TYPE UDT_MAN_CMD_WR :   // Manual commands from HMI
STRUCT
   CONV_Manual_ALL : BOOL;
   CONV_Man_ALL_FWD : BOOL;
   CONV_Man_ALL_REV : BOOL;
   M302M1_Manual : BOOL;
   M302M1_ManFWD : BOOL;
   M302M1_ManREV : BOOL;
   M302M1_ManSpeed : DINT;
   M302M2_Manual : BOOL;
   M302M2_ManFWD : BOOL;
   M302M2_ManREV : BOOL;
   M302M2_ManSpeed : DINT;
   M302M3_Manual : BOOL;
   M302M3_ManFWD : BOOL;
   M302M3_ManREV : BOOL;
   M302M3_ManSpeed : DINT;
   M302M4_Manual : BOOL;
   M302M4_ManFWD : BOOL;
   M302M4_ManREV : BOOL;
   M302M4_ManSpeed : DINT;
   M302M5_Manual : BOOL;
   M302M5_ManFWD : BOOL;
   M302M5_ManREV : BOOL;
   M302M5_ManSpeed : DINT;
   M302M6_Manual : BOOL;
   M302M6_ManFWD : BOOL;
   M302M6_ManREV : BOOL;
   M302M6_ManSpeed : DINT;
   M302M7_Manual : BOOL;
   M302M7_ManFWD : BOOL;
   M302M7_ManREV : BOOL;
   M302M7_ManSpeed : DINT;
   M303M1_Manual : BOOL;
   M303M1_ManFWD : BOOL;
   M303M1_ManREV : BOOL;
   M303M1_ManSpeed : DINT;
   M303M2_Manual : BOOL;
   M303M2_ManFWD : BOOL;
   M303M2_ManREV : BOOL;
   M303M2_ManSpeed : DINT;
   M304M1_Manual : BOOL;
   M304M1_ManFWD : BOOL;
   M304M1_ManREV : BOOL;
   M304M1_ManSpeed : DINT;
   M305M1_Manual : BOOL;
   M305M1_ManFWD : BOOL;
   M305M1_ManREV : BOOL;
   M305M1_ManSpeed : DINT;
   M306M1_Manual : BOOL;
   M306M1_ManFWD : BOOL;
   M306M1_ManREV : BOOL;
   M306M1_ManSpeed : DINT;
   M307AM1_Manual : BOOL;
   M307AM1_ManFWD : BOOL;
   M307AM1_ManREV : BOOL;
   M307AM1_ManSpeed : DINT;
   M307AM2_Manual : BOOL;
   M307AM2_ManFWD : BOOL;
   M307AM2_ManREV : BOOL;
   M307AM2_ManSpeed : DINT;
   M307AM3_Manual : BOOL;
   M307AM3_ManFWD : BOOL;
   M307AM3_ManREV : BOOL;
   M307AM3_ManSpeed : DINT;
   M307AM4_Manual : BOOL;
   M307AM4_ManFWD : BOOL;
   M307AM4_ManREV : BOOL;
   M307AM4_ManSpeed : DINT;
   M307BM1_Manual : BOOL;
   M307BM1_ManFWD : BOOL;
   M307BM1_ManREV : BOOL;
   M307BM1_ManSpeed : DINT;
   M307CM1_Manual : BOOL;
   M307CM1_ManFWD : BOOL;
   M307CM1_ManREV : BOOL;
   M307CM1_ManSpeed : DINT;
   M307DM1_Manual : BOOL;
   M307DM1_ManFWD : BOOL;
   M307DM1_ManREV : BOOL;
   M307DM1_ManSpeed : DINT;
   M307EM1_Manual : BOOL;
   M307EM1_ManFWD : BOOL;
   M307EM1_ManREV : BOOL;
   M307EM1_ManSpeed : DINT;
   M307FM1_Manual : BOOL;
   M307FM1_ManFWD : BOOL;
   M307FM1_ManREV : BOOL;
   M307FM1_ManSpeed : DINT;
   M310M1_Manual : BOOL;
   M310M1_ManFWD : BOOL;
   M310M1_ManREV : BOOL;
   M310M1_ManSpeed : DINT;
   M310M2_Manual : BOOL;
   M310M2_ManFWD : BOOL;
   M310M2_ManREV : BOOL;
   M310M2_ManSpeed : DINT;
   M310M3_Manual : BOOL;
   M310M3_ManFWD : BOOL;
   M310M3_ManREV : BOOL;
   M310M3_ManSpeed : DINT;
   M310M4_Manual : BOOL;
   M310M4_ManFWD : BOOL;
   M310M4_ManREV : BOOL;
   M310M4_ManSpeed : DINT;
   M310M5_Manual : BOOL;
   M310M5_ManFWD : BOOL;
   M310M5_ManREV : BOOL;
   M310M5_ManSpeed : DINT;
   M310M6_Manual : BOOL;
   M310M6_ManFWD : BOOL;
   M310M6_ManREV : BOOL;
   M310M6_ManSpeed : DINT;
   M310M7_Manual : BOOL;
   M310M7_ManFWD : BOOL;
   M310M7_ManREV : BOOL;
   M310M7_ManSpeed : DINT;
   M311M1_Manual : BOOL;
   M311M1_ManFWD : BOOL;
   M311M1_ManREV : BOOL;
   M311M1_ManSpeed : DINT;
   M311AM1_Manual : BOOL;
   M311AM1_ManFWD : BOOL;
   M311AM1_ManREV : BOOL;
   M311AM1_ManSpeed : DINT;
   M312M1_Manual : BOOL;
   M312M1_ManFWD : BOOL;
   M312M1_ManREV : BOOL;
   M312M1_ManSpeed : DINT;
   M312M2_Manual : BOOL;
   M312M2_ManFWD : BOOL;
   M312M2_ManREV : BOOL;
   M312M2_ManSpeed : DINT;
   M312M3_Manual : BOOL;
   M312M3_ManFWD : BOOL;
   M312M3_ManREV : BOOL;
   M312M3_ManSpeed : DINT;
   M315M1_Manual : BOOL;
   M315M1_ManFWD : BOOL;
   M315M1_ManREV : BOOL;
   M315M1_ManSpeed : DINT;
   M315M2_Manual : BOOL;
   M315M2_ManFWD : BOOL;
   M315M2_ManREV : BOOL;
   M315M2_ManSpeed : DINT;
   M315M3_Manual : BOOL;
   M315M3_ManFWD : BOOL;
   M315M3_ManREV : BOOL;
   M315M3_ManSpeed : DINT;
   M315M4_Manual : BOOL;
   M315M4_ManFWD : BOOL;
   M315M4_ManREV : BOOL;
   M315M4_ManSpeed : DINT;
   M315M5_Manual : BOOL;
   M315M5_ManFWD : BOOL;
   M315M5_ManREV : BOOL;
   M315M5_ManSpeed : DINT;
   M315M6_Manual : BOOL;
   M315M6_ManFWD : BOOL;
   M315M6_ManREV : BOOL;
   M315M6_ManSpeed : DINT;
   M315M7_Manual : BOOL;
   M315M7_ManFWD : BOOL;
   M315M7_ManREV : BOOL;
   M315M7_ManSpeed : DINT;
   M315AM1_Manual : BOOL;
   M315AM1_ManFWD : BOOL;
   M315AM1_ManREV : BOOL;
   M315AM1_ManSpeed : DINT;
   M316M1_Manual : BOOL;
   M316M1_ManFWD : BOOL;
   M316M1_ManREV : BOOL;
   M316M1_ManSpeed : DINT;
   M316AM1_Manual : BOOL;
   M316AM1_ManFWD : BOOL;
   M316AM1_ManREV : BOOL;
   M316AM1_ManSpeed : DINT;
   M317M1_Manual : BOOL;
   M317M1_ManFWD : BOOL;
   M317M1_ManREV : BOOL;
   M317M1_ManSpeed : DINT;
   M317M2_Manual : BOOL;
   M317M2_ManFWD : BOOL;
   M317M2_ManREV : BOOL;
   M317M2_ManSpeed : DINT;
   M317M3_Manual : BOOL;
   M317M3_ManFWD : BOOL;
   M317M3_ManREV : BOOL;
   M317M3_ManSpeed : DINT;
   M350M1_Manual : BOOL;
   M350M1_ManFWD : BOOL;
   M350M1_ManREV : BOOL;
   M350M1_ManSpeed : DINT;
   M351M1_Manual : BOOL;
   M351M1_ManFWD : BOOL;
   M351M1_ManREV : BOOL;
   M351M1_ManSpeed : DINT;
   M360M1_Manual : BOOL;
   M360M1_ManFWD : BOOL;
   M360M1_ManREV : BOOL;
   M360M1_ManSpeed : DINT;
END_STRUCT
END_TYPE

TYPE UDT_MOTOR_HMR :
STRUCT
   M302M1_Feedback : BOOL;
   M302M1_Faulted : BOOL;
   M302M1_FaultCode : DINT;
   M302M1_OutSpeed : DINT;
   M302M1_OutCurrent : DINT;
   M302M2_Feedback : BOOL;
   M302M2_Faulted : BOOL;
   M302M2_FaultCode : DINT;
   M302M2_OutSpeed : DINT;
   M302M2_OutCurrent : DINT;
   M302M3_Feedback : BOOL;
   M302M3_Faulted : BOOL;
   M302M3_FaultCode : DINT;
   M302M3_OutSpeed : DINT;
   M302M3_OutCurrent : DINT;
   M302M4_Feedback : BOOL;
   M302M4_Faulted : BOOL;
   M302M4_FaultCode : DINT;
   M302M4_OutSpeed : DINT;
   M302M4_OutCurrent : DINT;
   M302M5_Feedback : BOOL;
   M302M5_Faulted : BOOL;
   M302M5_FaultCode : DINT;
   M302M5_OutSpeed : DINT;
   M302M5_OutCurrent : DINT;
   M302M6_Feedback : BOOL;
   M302M6_Faulted : BOOL;
   M302M6_FaultCode : DINT;
   M302M6_OutSpeed : DINT;
   M302M6_OutCurrent : DINT;
   M302M7_Feedback : BOOL;
   M302M7_Faulted : BOOL;
   M302M7_FaultCode : DINT;
   M302M7_OutSpeed : DINT;
   M302M7_OutCurrent : DINT;
   M303M1_Feedback : BOOL;
   M303M1_Faulted : BOOL;
   M303M1_FaultCode : DINT;
   M303M1_OutSpeed : DINT;
   M303M1_OutCurrent : DINT;
   M303M2_Feedback : BOOL;
   M303M2_Faulted : BOOL;
   M303M2_FaultCode : DINT;
   M303M2_OutSpeed : DINT;
   M303M2_OutCurrent : DINT;
   M304M1_Feedback : BOOL;
   M304M1_Faulted : BOOL;
   M304M1_FaultCode : DINT;
   M304M1_OutSpeed : DINT;
   M304M1_OutCurrent : DINT;
   M305M1_Feedback : BOOL;
   M305M1_Faulted : BOOL;
   M305M1_FaultCode : DINT;
   M305M1_OutSpeed : DINT;
   M305M1_OutCurrent : DINT;
   M306M1_Feedback : BOOL;
   M306M1_Faulted : BOOL;
   M306M1_FaultCode : DINT;
   M306M1_OutSpeed : DINT;
   M306M1_OutCurrent : DINT;
   M307AM1_Feedback : BOOL;
   M307AM1_Faulted : BOOL;
   M307AM1_FaultCode : DINT;
   M307AM1_OutSpeed : DINT;
   M307AM1_OutCurrent : DINT;
   M307AM2_Feedback : BOOL;
   M307AM2_Faulted : BOOL;
   M307AM2_FaultCode : DINT;
   M307AM2_OutSpeed : DINT;
   M307AM2_OutCurrent : DINT;
   M307AM3_Feedback : BOOL;
   M307AM3_Faulted : BOOL;
   M307AM3_FaultCode : DINT;
   M307AM3_OutSpeed : DINT;
   M307AM3_OutCurrent : DINT;
   M307AM4_Feedback : BOOL;
   M307AM4_Faulted : BOOL;
   M307AM4_FaultCode : DINT;
   M307AM4_OutSpeed : DINT;
   M307AM4_OutCurrent : DINT;
   M307BM1_Feedback : BOOL;
   M307BM1_Faulted : BOOL;
   M307BM1_FaultCode : DINT;
   M307BM1_OutSpeed : DINT;
   M307BM1_OutCurrent : DINT;
   M307CM1_Feedback : BOOL;
   M307CM1_Faulted : BOOL;
   M307CM1_FaultCode : DINT;
   M307CM1_OutSpeed : DINT;
   M307CM1_OutCurrent : DINT;
   M307DM1_Feedback : BOOL;
   M307DM1_Faulted : BOOL;
   M307DM1_FaultCode : DINT;
   M307DM1_OutSpeed : DINT;
   M307DM1_OutCurrent : DINT;
   M307EM1_Feedback : BOOL;
   M307EM1_Faulted : BOOL;
   M307EM1_FaultCode : DINT;
   M307EM1_OutSpeed : DINT;
   M307EM1_OutCurrent : DINT;
   M307FM1_Feedback : BOOL;
   M307FM1_Faulted : BOOL;
   M307FM1_FaultCode : DINT;
   M307FM1_OutSpeed : DINT;
   M307FM1_OutCurrent : DINT;
   M310M1_Feedback : BOOL;
   M310M1_Faulted : BOOL;
   M310M1_FaultCode : DINT;
   M310M1_OutSpeed : DINT;
   M310M1_OutCurrent : DINT;
   M310M2_Feedback : BOOL;
   M310M2_Faulted : BOOL;
   M310M2_FaultCode : DINT;
   M310M2_OutSpeed : DINT;
   M310M2_OutCurrent : DINT;
   M310M3_Feedback : BOOL;
   M310M3_Faulted : BOOL;
   M310M3_FaultCode : DINT;
   M310M3_OutSpeed : DINT;
   M310M3_OutCurrent : DINT;
   M310M4_Feedback : BOOL;
   M310M4_Faulted : BOOL;
   M310M4_FaultCode : DINT;
   M310M4_OutSpeed : DINT;
   M310M4_OutCurrent : DINT;
   M310M5_Feedback : BOOL;
   M310M5_Faulted : BOOL;
   M310M5_FaultCode : DINT;
   M310M5_OutSpeed : DINT;
   M310M5_OutCurrent : DINT;
   M310M6_Feedback : BOOL;
   M310M6_Faulted : BOOL;
   M310M6_FaultCode : DINT;
   M310M6_OutSpeed : DINT;
   M310M6_OutCurrent : DINT;
   M310M7_Feedback : BOOL;
   M310M7_Faulted : BOOL;
   M310M7_FaultCode : DINT;
   M310M7_OutSpeed : DINT;
   M310M7_OutCurrent : DINT;
   M311M1_Feedback : BOOL;
   M311M1_Faulted : BOOL;
   M311M1_FaultCode : DINT;
   M311M1_OutSpeed : DINT;
   M311M1_OutCurrent : DINT;
   M311AM1_Feedback : BOOL;
   M311AM1_Faulted : BOOL;
   M311AM1_FaultCode : DINT;
   M311AM1_OutSpeed : DINT;
   M311AM1_OutCurrent : DINT;
   M312M1_Feedback : BOOL;
   M312M1_Faulted : BOOL;
   M312M1_FaultCode : DINT;
   M312M1_OutSpeed : DINT;
   M312M1_OutCurrent : DINT;
   M312M2_Feedback : BOOL;
   M312M2_Faulted : BOOL;
   M312M2_FaultCode : DINT;
   M312M2_OutSpeed : DINT;
   M312M2_OutCurrent : DINT;
   M312M3_Feedback : BOOL;
   M312M3_Faulted : BOOL;
   M312M3_FaultCode : DINT;
   M312M3_OutSpeed : DINT;
   M312M3_OutCurrent : DINT;
   M315M1_Feedback : BOOL;
   M315M1_Faulted : BOOL;
   M315M1_FaultCode : DINT;
   M315M1_OutSpeed : DINT;
   M315M1_OutCurrent : DINT;
   M315M2_Feedback : BOOL;
   M315M2_Faulted : BOOL;
   M315M2_FaultCode : DINT;
   M315M2_OutSpeed : DINT;
   M315M2_OutCurrent : DINT;
   M315M3_Feedback : BOOL;
   M315M3_Faulted : BOOL;
   M315M3_FaultCode : DINT;
   M315M3_OutSpeed : DINT;
   M315M3_OutCurrent : DINT;
   M315M4_Feedback : BOOL;
   M315M4_Faulted : BOOL;
   M315M4_FaultCode : DINT;
   M315M4_OutSpeed : DINT;
   M315M4_OutCurrent : DINT;
   M315M5_Feedback : BOOL;
   M315M5_Faulted : BOOL;
   M315M5_FaultCode : DINT;
   M315M5_OutSpeed : DINT;
   M315M5_OutCurrent : DINT;
   M315M6_Feedback : BOOL;
   M315M6_Faulted : BOOL;
   M315M6_FaultCode : DINT;
   M315M6_OutSpeed : DINT;
   M315M6_OutCurrent : DINT;
   M315M7_Feedback : BOOL;
   M315M7_Faulted : BOOL;
   M315M7_FaultCode : DINT;
   M315M7_OutSpeed : DINT;
   M315M7_OutCurrent : DINT;
   M315AM1_Feedback : BOOL;
   M315AM1_Faulted : BOOL;
   M315AM1_FaultCode : DINT;
   M315AM1_OutSpeed : DINT;
   M315AM1_OutCurrent : DINT;
   M316M1_Feedback : BOOL;
   M316M1_Faulted : BOOL;
   M316M1_FaultCode : DINT;
   M316M1_OutSpeed : DINT;
   M316M1_OutCurrent : DINT;
   M316AM1_Feedback : BOOL;
   M316AM1_Faulted : BOOL;
   M316AM1_FaultCode : DINT;
   M316AM1_OutSpeed : DINT;
   M316AM1_OutCurrent : DINT;
   M317M1_Feedback : BOOL;
   M317M1_Faulted : BOOL;
   M317M1_FaultCode : DINT;
   M317M1_OutSpeed : DINT;
   M317M1_OutCurrent : DINT;
   M317M2_Feedback : BOOL;
   M317M2_Faulted : BOOL;
   M317M2_FaultCode : DINT;
   M317M2_OutSpeed : DINT;
   M317M2_OutCurrent : DINT;
   M317M3_Feedback : BOOL;
   M317M3_Faulted : BOOL;
   M317M3_FaultCode : DINT;
   M317M3_OutSpeed : DINT;
   M317M3_OutCurrent : DINT;
   M350M1_Feedback : BOOL;
   M350M1_Faulted : BOOL;
   M350M1_FaultCode : DINT;
   M350M1_OutSpeed : DINT;
   M350M1_OutCurrent : DINT;
   M351M1_Feedback : BOOL;
   M351M1_Faulted : BOOL;
   M351M1_FaultCode : DINT;
   M351M1_OutSpeed : DINT;
   M351M1_OutCurrent : DINT;
   M360M1_Feedback : BOOL;
   M360M1_Faulted : BOOL;
   M360M1_FaultCode : DINT;
   M360M1_OutSpeed : DINT;
   M360M1_OutCurrent : DINT;
END_STRUCT
END_TYPE

TYPE UDT_PLANT_CONSTANTS :
STRUCT
   dPLC_ID : DINT;   // 1= PLC#1 2= PLC#2
   dOP_Side : DINT;   // 0=Operator side right; 1=Operator side left
   dZ1ConveyorNumber : DINT;   // Conveyor number in Z301
   dZ1TotalLength_cmm : DINT;   // Z301 total length of tracking [mm/100]
   dZ2ConveyorNumber : DINT;   // Conveyor number in Z302
   dZ2TotalLength_cmm : DINT;   // Z302 total length of tracking [mm/100]
   dZ3ConveyorNumber : DINT;   // Conveyor number in Z303
   dZ3TotalLength_cmm : DINT;   // Z303 total length of tracking [mm/100]
   dTrimDeckNumber : DINT;   // Trimming deck number
   dTrimWheelsNumber : DINT;   // Trimming wheels number
   dSplitBarNumber : DINT;   // Split bar number
   dSepRollNumber : DINT;   // Separator roll number
   dTrackWindows_cmm : DINT;   // Tracking windows step [mm/100]
   dMaxScanSpace_cmm : DINT;   // Max space calculated on each scan at maximum line speed [mm/100]
   rgdAccDecRamps : REAL[4];   // Acceleration / Deceleration ramps used in main line [m/s2]
   dMaxLineSpeed_mm_min : DINT;   // Max line speed [mm/min]
   dMinLineSpeed_mm_min : DINT;   // Min line speed [mm/min]
   dMaxLineSnapSpeed_mm_min : DINT;   // Max line speed for snapping area [mm/min]
   dMinLineSnapSpeed_mm_min : DINT;   // Min line speed for snapping area [mm/min]
   dMaxLehrSpeed_mm_min : DINT;   // Max lehr speed [mm/min]
   dMinLehrSpeed_mm_min : DINT;   // Min lehr speed [mm/min]
   rMaxSpeedRatio : REAL;   // Max speed ratio [Num]
   rMinSpeedRatio : REAL;   // Min speed ratio [Num]
   rMaxSpeedSnapRatio : REAL;   // Max speed ratio for snapping area [Num]
   rMinSpeedSnapRatio : REAL;   // Min speed ratio for snapping area [Num]
   dZ1CleaningSpeed_mm_min : DINT;   // Cleaning speed Z301 [mm/min] (Optional if no cooling on motors)
   dMaxNumPlates : DINT;   // Maximum number of plates in tracking (circular buffer positions)
   dMaxNumHeadTail : DINT;   // Maximum number of head tail
   rgdLiteLimits_cmm : DINT[20];   // Lite limits [mm/100] (Length,width...)
   rgdCapLimits_cmm : DINT[5];   // Cap limits [mm/100] (Length,width,max num lites,...)
   rgdConvoyLimits_cmm : DINT[5];   // Convoy limits [mm/100] (Length,width,max num caps,...)
   rgdRibbonLimits_cmm : DINT[5];   // Ribbon limits [mm/100]
   rgdWanderLimits : DINT[2];   // Wander limits [mm/100]
   dNumOfConveyors : DINT;   // Number of conveyors [Num]
   dNumCapsConveyor : DINT;   // Number of caps per conveyor [Num]
   dNumCapsMaxConvoy : DINT;   // Maximum number of caps per convoy [Num]
   dNumLitesMaxCap : DINT;   // Maximum number of lites per cap [Num]
   dNumPlateSearch : DINT;   // Number of plates to search in Search function [Num]
   dNumOfUnloadDestinations : DINT;   // Number of possible destinations for stack [Num]
END_STRUCT
END_TYPE

TYPE UDT_PlateData_Convoy :
STRUCT
   dSyncHead : DINT;   // Synchro Head
   dIDTx : DINT;
   dTotLenght_cmm : DINT;
   dTotWidth_cmm : DINT;
   dFormat : DINT;   // 1=JS 2=LES, 3=SSS
   dNumLites : DINT;   // Num Lite on board
   dPositionLite : DINT;   // 0=Centre Line, 1=Right Side Line. 2 Left Side Line
   tLite : UDT_PlateData_Convoy_Lite[2];
   dSyncTail : DINT;   // Synchro Tail
END_STRUCT
END_TYPE

TYPE UDT_PlateData_Convoy_Lite :
STRUCT
   dID : DINT;   // ID lite
   dProduction_ID : DINT;   // ID Production
   dLenght_cmm : DINT;   // Lenght Lite
   dWidth_cmm : DINT;   // Width Lite
   dThick_cmm : DINT;   // Thickness Lite
   rgxOrigin : DINT;   // Origin plate
   rgxMain : DINT;   // Main destination plate
   rgxAlternative : DINT;   // Alternative destination plate
   xCoated : BOOL;   // Type Coated
   xCoverPlate : BOOL;   // Type Cover
END_STRUCT
END_TYPE

TYPE UDT_SearchPlateAuxData :   // Auxiliary data for searching plate
STRUCT
   dIDMemory : DINT;   // ID Memory
   dReaction_cmm : DINT;   // Reation space [mm/100]
   dPositionDecision_cmm : DINT;   // Decision position [mm/100]
   dPositionStopSearch_cmm : DINT;   // Stop search position [mm/100]
   dPositionStopHooked_cmm : DINT;   // Stop hooked position [mm/100]
   dIndex : DINT;   // Index
   xIndexCons : BOOL;   // Index consistent
   xPlateHooked : BOOL;   // Plate hooked
   OS_xPlateInWindows : BOOL;   // OS Plate in windows
   OF_xPlateInWindows : BOOL;   // OF Plate in windows
   OSR_xPlateInWindows : BOOL;   // OSR Plate in windows
   OSF_xPlateInWindows : BOOL;   // OSF Plate in windows
   OSR_xPlateOutHooked : BOOL;   // OSR Plate hooked
   OS_xPlateOutHooked : BOOL;   // OS Plate hooked
   tResult : GP_TrackingSearchPlate_STC;   // Search plate data result
END_STRUCT
END_TYPE

TYPE UDT_StandConv :
STRUCT
   ST_rgxRampInProgress : DINT;   // Ramp in progress
   ST_rgxDecInProgress : DINT;   // Deceleration in progress
   ST_rgxAccInProgress : DINT;   // Acceleration in progress
   ST_rgxBrakeRelease : DINT;   // Brake release
   ST_rgxBrakeFeedback : DINT;   // Brake feedback
   ST_rgxConveyorOutRunSgm : DINT;   // Single motor conveyor out run
   ST_rgxOutMotorRunSgm : DINT;   // Single motor out run active
   ST_xDriveInDec : BOOL;   // At least one drive in deceleration
   ST_xPositionReached : BOOL;   // Position reached
   ST_xManualCmdEnabled : BOOL;   // Manual command enabled
   ST_xEnableControlError : BOOL;   // Enable control error
   ST_xRotationFeedback : BOOL;   // Rotation feedback
   ST_xCleaningConditionOK : BOOL;   // Cleaning condition OK
   ST_xCleaningEnabled : BOOL;   // Cleaning enabled
   ST_xReqCleaning : BOOL;   // Cleaning request
   ST_xOutputEnable : BOOL;   // Output enable
   ST_xFaulted : BOOL;   // Conveyor faulted
   ST_xStopMachineFault : BOOL;   // Stopped machine faults
   ST_xStopNextCycleFault : BOOL;   // Stopped next cycle faults
   ST_xWarningFault : BOOL;   // Warning fault
   ST_xStopCycleConditionOK : BOOL;   // Condition OK for stop cycle
   ST_xConveyorOutRun : BOOL;   // Conveyor out run
   ST_xOutMotorRun : BOOL;   // Motor out run active
   ST_xStopConveyorDuringClean : BOOL;   // Stop conveyor during cleaning
   ST_xStopConveyor : BOOL;   // Stop conveyor
   ST_xStopConveyorM1 : BOOL;   // Stop conveyor M1
   ST_xStopConveyorM2 : BOOL;   // Stop conveyor M2
   ST_xStopPlateAtEndConveyor : BOOL;   // Stop plate at end of conveyor
   ST_xAxleReadyToMoveDelayed : BOOL;   // Axle ready to move delayed
   ST_xSafetyConveyor : BOOL;   // Safety conveyor
   ST_xOneReqActive : BOOL;   // At least one request active
   ST_xPositionReqActive : BOOL;   // Positioning request active
   ST_xPositionReqActiveM1 : BOOL;   // Positioning request active M1
   ST_xPositionReqActiveM2 : BOOL;   // Positioning request active M2
   ST_xStopEndConveyorReached : BOOL;   // Stop at end of conveyor reached
   ST_xWaitFeedbackRestart : BOOL;   // Wait feedback restart
   ST_xWaitStopConveyor : BOOL;   // Wait stop conveyor
   ST_xInitialCondition : BOOL;   // Only for optimize external decision
   ST_xRestartActive : BOOL;   // Conveyor Restart Active
   xReqStop : BOOL;   // Request stop
   xReqStopEndConveyor : BOOL;   // Request stop at end of conveyor
   xReqBypassEndStop : BOOL;   // Request bypass end stop
   xReqStopNextConveyor : BOOL;   // Request stop next conveyor
   xReqStopM1 : BOOL;   // Request stop motor M1
   xReqStopM2 : BOOL;   // Request stop motor M2
   xReqBypassEndConveyorM1 : BOOL;   // Request bypass end conveyor M1
   xReqBypassEndConveyorM2 : BOOL;   // Request bypass end conveyor M2
   xReqPositioningHead : BOOL;   // Request positioning with photocell on head
   xReqPositioningTail : BOOL;   // Request positioning with photocell on tail
   xReqPositioningAbs : BOOL;   // Request absolute positioning
   xReqPositioningHeadM1 : BOOL;   // Request positioning with photocell on head M1
   xReqPositioningTailM1 : BOOL;   // Request positioning with photocell on tail M1
   xReqPositioningAbsM1 : BOOL;   // Request absolute positioning M1
   xReqPositioningHeadM2 : BOOL;   // Request positioning with photocell on head M2
   xReqPositioningTailM2 : BOOL;   // Request positioning with photocell on tail M2
   xReqPositioningAbsM2 : BOOL;   // Request absolute positioning M2
   xReqSpeed : BOOL;   // Request speed
   xReqExtStopLoadNewPlate : BOOL;   // Request external condition stop load new plate
   OS_xExpTimeOutAnomaly : BOOL;   // OS Expired timeout anomaly
   OS_xRunMotor : BOOL;   // OS Run motor
   OSF_xCleaningAccZone : BOOL;   // OSF Cleaning acceleration zone
   OSR_xCleaningAccZone : BOOL;   // OSR Cleaning acceleration zone
   OSF_xCleaningZoneAcc : BOOL;   // OSF Cleaning zone acceleration
   OSR_xRunMotor : BOOL;   // OSR Run motor
   OSR_xWaitStop : BOOL;   // OSR Wait stop
   OS_xStartCount : DINT;   // OS Start count positioning
   OSR_xStartCount : DINT;   // OSR Start count positioning
   INPUT_xPowerModuleON : BOOL;   // Power module ON
   INPUT_xSafetyConveyor : BOOL;   // Safety conveyor
   INPUT_xSpeedRequest : BOOL;   // Speed request
   INPUT_xPhotocellPositioning : DINT;   // Photocell positioning
   INPUT_xBrakingResistor : DINT;   // Braking Resistor
   INPUT_xDriveInhibit : DINT;   // Drive inhibit
   INPUT_xDriveReady : DINT;   // Drive ready
   INPUT_xDriveError : DINT;   // Drive Error
   INPUT_xDriveFeedback : DINT;   // Drive Feedback
   INPUT_xDriveDeceleration : DINT;   // Drive deceleration
   INPUT_xDriveAcceleration : DINT;   // Drive acceleration
   INPUT_xLocalSafetySwitch : DINT;   // Local Safety Switch
   INPUT_xMotorThermalProbe : DINT;   // Motor Thermal Probe
   INPUT_xProtectionMotor : DINT;   // Protection Motor
   INPUT_xProtectionCoolingFan : DINT;   // Protection cooling fan
   INPUT_xFeedbackCoolingFan : DINT;   // Feedback cooling fan
   INPUT_xDrivePositionReached : DINT;   // Drive position reached
   INPUT_rgdRefSpeed_mm_min : DINT[5];   // Reference speed (0=AutoSpeed, 1=LehrSpeed, 2=CleaningSpeed, 3=SpecialSpeed, 4=ManualSpeed) [mm/min]
   INPUT_dIndexSpeedReq : DINT;   // Use together request special speed
   tIN_Zone : UDT_IN_Zone;   // Zone inputs
   OUTPUT_xDriveReset : DINT;   // Drive reset faults
   OUTPUT_xDriveEnable : DINT;   // Output
   OUTPUT_xRun : DINT;   // Run
   OUTPUT_xReverse : DINT;   // Reverse
   OUTPUT_xPositioning : DINT;   // Positioning
   OUTPUT_xChangeSpeed : DINT;   // Change speed
   AUX_rgdCurrentSpeed_mm_min : DINT[2];   // Conveyor current speed [mm/min]
   AUX_rgdRequestSpeed_mm_min : DINT[2];   // Conveyor requested speed [mm/min]
   AUX_rgdLastIDPlateLoaded : DINT[2];   // Last ID plate loaded
   AUX_rgdLoadPreset_cmm : DINT[2];   // Load preset quote [mm/100]
   AUX_rgdLoadPresetWithRestart_cmm : DINT[2];   // Load preset quote in case of restart active [mm/100]
   AUX_rgdAccSpace_cmm : DINT[2];   // Acceleration space [mm/100]
   AUX_rgdDecSpace_cmm : DINT[2];   // Deceleration space [mm/100]
   AUX_rgdTarget_cmm : DINT[2];   // Positioning target [mm/100]
   AUX_rgdStepAdvancement_cmm : DINT[2];   // Step space per scan [mm/100]
   AUX_rgrAcc_m_s2 : REAL[2];   // Acceleration ramp [m/s2]
   AUX_rgrDec_m_s2 : REAL[2];   // Deceleration ramp [m/s2]
   AUX_rgrReminderStep : REAL[2];   // Reminder Step [ms]
   AUX_rgrSpeedIncrement_mm_min : REAL[2];   // Head position [mm/min]
   AUX_rgrCurrentDriveSpeed_mm_min : REAL[2];   // Drive current speed [mm/min]
   tmOFF_DriveEnable : TIMER[2];   // Drive enable timer
   tmON_DelayReadyToMove : TIMER[2];   // Delay timer for ready to move
   tmON_FeedbackDriveReady : TIMER[2];   // Drive ready feedback timer
   tmON_FeedbackTimeout : TIMER[2];   // Feedback timeout
   tmOFF_DelayPhotocellTail : TIMER[2];   // Delay timer for tail photocell
   tmON_PhFilter : TIMER[2];   // Start count photocell filter
   tmON_EnableActivedFilter : TIMER[2];   // Filter on enable timer
END_STRUCT
END_TYPE

TYPE UDT_Tracking :
STRUCT
   dPosition_cmm : DINT;   // Barycenter tracking position from snapbar [cmm]
   dPositionHead_cmm : DINT;   // Head tracking position from snapbar [cmm]
   dPositionTail_cmm : DINT;   // Tail tracking position from snapbar [cmm]
   dPreviousCapIndex : DINT;   // Previous cap index data (if Next & Previous are null -> No convoy) [Num]
   dNextCapIndex : DINT;   // Next cap index data (if Next & Previous are null -> No convoy) [Num]
   dLength_cmm : DINT;   // Cap Length [cmm]
   dLengthConvoy : DINT;   // Convoy Length [cmm]
   dGapConvoy : DINT;   // Gap Convoy [cmm]
   dIndexConvHead : DINT;   // Index conveyor head [Num]
   dIndexCapInConvHead : DINT;   // Index cap inside conveyor head [Num]
   dIndexConvTail : DINT;   // Index conveyor tail [Num]
   dIndexCapInConvTail : DINT;   // Index cap inside conveyor head [Num]
   dIndexMotorStepAdv : DINT;   // Index motor used for advancement [Motor1:0,Motor2:1]
   dIndexConvNotCons : DINT;   // Reserved. Index of conveyor not considered in tracking for speed
   dLastConv : DINT;   // Reserved. Last conveyor plate presence
   dLastConvTail : DINT;   // Reserved. Last conveyor plate presence tail
   xNotConsConvTrk : BOOL;   // Reserved. Not considered in the conveyor presence
   xHoldAdvancement : BOOL;   // Hold tracking plate
   xNotShownInScada : BOOL;   // Not shown in scada system
   xFirstPlateConvoy : BOOL;   // First plate of the convoy
   xLastPlateConvoy : BOOL;   // Last plate of the convoy
   xPlateInConvoy : BOOL;   // Plate in the middle of convoy
END_STRUCT
END_TYPE

TYPE WorkingFlags_Conveyor :
STRUCT
   xReqStop : BOOL;   // Request stop of conveyor
   xBypassReqEndStop : BOOL;   // Request bypass stop at end of conveyor
   xReqStopEndConveyor : BOOL;   // Request stop at end of conveyor
   xReqStopM1 : BOOL;   // Request stop motor M1
   xReqStopM2 : BOOL;   // Request stop motor M2
   xReqPositioningHead : BOOL;   // Request infinite positioning on head (Using positioner target)
   xReqPositioningTail : BOOL;   // Request infinite positioning on tail (Using positioner target)
   xReqPositioningAbs : BOOL;   // Request absolute positioning (Using positioner target)
   xDoneStop : BOOL;   // Done stop of conveyor
   xDoneBypassEndStop : BOOL;   // Done bypass stop at end of conveyor
   xDoneStopEndConveyor : BOOL;   // Done stop at end of conveyor
   xDoneStopM1 : BOOL;   // Done stop of motor M1
   xDoneStopM2 : BOOL;   // Done stop of motor M2
   xDoneHeadPositioning : BOOL;   // Done infinite positioning on head (Using positioner target)
   xDoneTailPositioning : BOOL;   // Done infinite positioning on tail (Using positioner target)
   xDoneAbsPositioning : BOOL;   // Done absolute positioning (Using positioner target)
   dTarget_cmm : DINT;   // Target [mm/100]
   dSpare0 : DINT;   // Spare
   dSpare1 : DINT;   // Spare
   dSpare2 : DINT;   // Spare
   dSpare3 : DINT;   // Spare
END_STRUCT
END_TYPE

TYPE WorkingFlags_GeomCamera :
STRUCT
   xReqIspection : BOOL;   // Request ispection
   xDoneIspection : BOOL;   // Done ispection
END_STRUCT
END_TYPE

TYPE WorkingFlags_Powder :
STRUCT
   xReqPowderA : BOOL;   // Request powder type A
   xReqPowderB : BOOL;   // Request powder type B
   xDonePowderA : BOOL;   // Done powder type A
   xDonePowderB : BOOL;   // Done powder type B
END_STRUCT
END_TYPE

TYPE WorkingFlags_Rotator :
STRUCT
   xReqRotationCw : BOOL;   // Request clockwise rotation
   xReqRotationCcw : BOOL;   // Request counterclockwise rotation
   xDoneRotationCw : BOOL;   // Done clockwise rotation
   xDoneRotationCcw : BOOL;   // Done counterclockwise rotation
   dStepNumb : DINT;   // Number of steps in rotation (0=90° 1=180° 2=270°)
END_STRUCT
END_TYPE

TYPE WorkingFlags_Selvedge :
STRUCT
   dReqTrim3OpSide : DINT;   // Request Trim 3 Op. Side (Triple edge) with trim wheel number [x=Num]
   dReqTrim2OpSide : DINT;   // Request Trim 2 Op. Side (Double edge) with trim wheel number [x=Num]
   dReqTrim1OpSide : DINT;   // Request Trim 1 Op. Side (Single edge) with trim wheel number [x=Num]
   dReqTrim1OppOpSide : DINT;   // Request Trim 1 Oppo. Op. Side (Single edge) with trim wheel number [x=Num]
   dReqTrim2OppOpSide : DINT;   // Request Trim 2 Oppo. Op. Side (Double edge) with trim wheel number [x=Num]
   dReqTrim3OppOpSide : DINT;   // Request Trim 3 Oppo. Op. Side (Triple edge) with trim wheel number [x=Num]
   dDoneTrim3OpSide : DINT;   // Done Trim 3 Op. Side (Triple edge) with trim wheel number [x=Num]
   dDoneTrim2OpSide : DINT;   // Done Trim 2 Op. Side (Double edge) with trim wheel number [x=Num]
   dDoneTrim1OpSide : DINT;   // Done Trim 1 Op. Side (Single edge) with trim wheel number [x=Num]
   dDoneTrim1OppOpSide : DINT;   // Done Trim 1 Oppo. Op. Side (Single edge) with trim wheel number [x=Num]
   dDoneTrim2OppOpSide : DINT;   // Done Trim 2 Oppo. Op. Side (Double edge) with trim wheel number [x=Num]
   dDoneTrim3OppOpSide : DINT;   // Done Trim 3 Oppo. Op. Side (Triple edge) with trim wheel number [x=Num]
   dFramePositionSelectionOpSide_cmm : DINT;   // Translation position of frame on operator side [mm/100]
   dFramePositionSelectionOppOpSide_cmm : DINT;   // Translation position of frame on opposite operator side [mm/100]
END_STRUCT
END_TYPE

ADD_ON_INSTRUCTION GP_AccessArea   (* revision 1.0 *)
VAR_IN_OUT
   STC : GP_AccessArea_STC; {required}
END_VAR
VAR_INPUT
   IN_xAccSelector : BOOL; {access None, required}
   IN_xAccButton : BOOL; {access None, required}
   IN_xConditionOkAccess : BOOL; {access None, required}
   IN_xConditionOkForcedAccess : BOOL; {access None, required}
   IN_xLampClock : BOOL; {access None, required}
END_VAR
VAR_OUTPUT
   OUT_xOpeningDoor : BOOL; {access None}
   OUT_xLamp : BOOL; {access None, required}
END_VAR

ROUTINE Logic   (* ladder *)
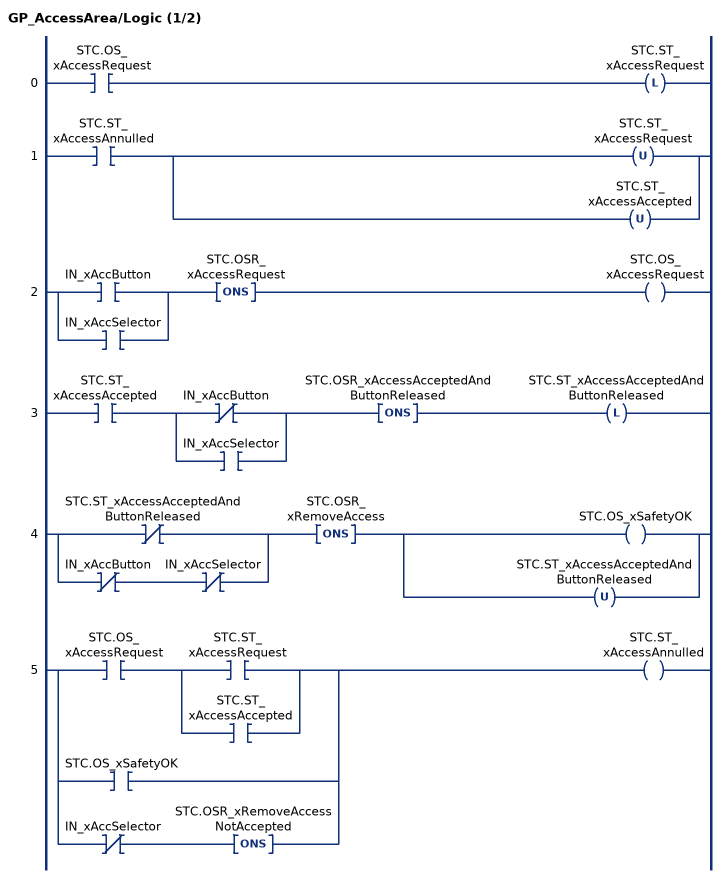
   0: XIC(STC.OS_xAccessRequest)OTL(STC.ST_xAccessRequest);
   1: XIC(STC.ST_xAccessAnnulled)[OTU(STC.ST_xAccessRequest) ,OTU(STC.ST_xAccessAccepted) ];
   2: [XIC(IN_xAccButton) ,XIC(IN_xAccSelector) ]ONS(STC.OSR_xAccessRequest)OTE(STC.OS_xAccessRequest);
   3: XIC(STC.ST_xAccessAccepted)[XIO(IN_xAccButton) ,XIC(IN_xAccSelector) ]ONS(STC.OSR_xAccessAcceptedAndButtonReleased)OTL(STC.ST_xAccessAcceptedAndButtonReleased);
   4: [XIO(STC.ST_xAccessAcceptedAndButtonReleased) ,XIO(IN_xAccButton) XIO(IN_xAccSelector) ]ONS(STC.OSR_xRemoveAccess)[OTE(STC.OS_xSafetyOK) ,OTU(STC.ST_xAccessAcceptedAndButtonReleased) ];
   5: [XIC(STC.OS_xAccessRequest) [XIC(STC.ST_xAccessRequest) ,XIC(STC.ST_xAccessAccepted) ] ,XIC(STC.OS_xSafetyOK) ,XIO(IN_xAccSelector) ONS(STC.OSR_xRemoveAccessNotAccepted) ]OTE(STC.ST_xAccessAnnulled);
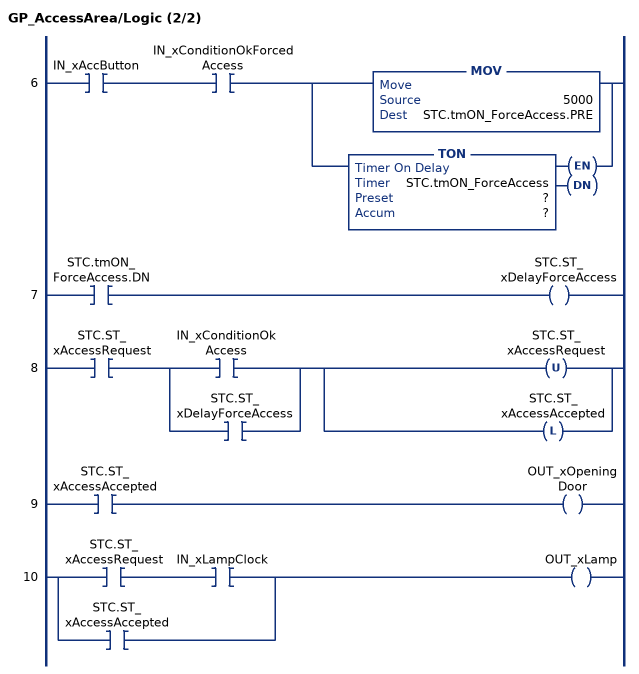
   6: XIC(IN_xAccButton)XIC(IN_xConditionOkForcedAccess)[MOV(5000,STC.tmON_ForceAccess.PRE) ,TON(STC.tmON_ForceAccess,?,?) ];
   7: XIC(STC.tmON_ForceAccess.DN)OTE(STC.ST_xDelayForceAccess);
   8: XIC(STC.ST_xAccessRequest)[XIC(IN_xConditionOkAccess) ,XIC(STC.ST_xDelayForceAccess) ][OTU(STC.ST_xAccessRequest) ,OTL(STC.ST_xAccessAccepted) ];
   9: XIC(STC.ST_xAccessAccepted)OTE(OUT_xOpeningDoor);
   10: [XIC(STC.ST_xAccessRequest) XIC(IN_xLampClock) ,XIC(STC.ST_xAccessAccepted) ]OTE(OUT_xLamp);
END_ROUTINE
END_ADD_ON_INSTRUCTION
